(* Logix 5000 project; controller WED2413001_BI600_AB vendor 1 type 14 code 192 rev 35.11; software revision 35.01 *)
// WED2413001_BI600_AB- automatically dispenses film on a roll, cuts, seals and inserts bags into cases, trays and bins

TASK MainTask (continuous, watchdog 500 ms) : BI600_MainProgram

MODULES
   Local : vendor 1 type 14 code 192 (5069 0, rev 35.11)
      VFD1_FILM_UNWIND : PowerFlex 525-EENET (Ethernet 192.168.5.38, rev 7.1, Output RPI 20 ms)   // PowerFlex 525 AC Drive, with Embedded EtherNet/IP and Safety, 200...240V AC, 3 Phase, 5.0 Amps, 1 H
      Cuffer_servo_UpDown : vendor 1 type 37 code 73 (Ethernet 192.168.5.30, rev 13.1, A_MotionDiagnostics RPI 1 ms, B_MotionSync RPI 1 ms)   // ALLEN BRADLEY 2198-C1015-ERS KINETIX 5300 SERVO VARIATEUR, 1.5KW 200V
      Cuffer_servomotor_OpenClose : 2198-C1004-ERS (Ethernet 192.168.5.31, rev 13.1, A_MotionDiagnostics RPI 1 ms, B_MotionSync RPI 1 ms)   // KINETIX 5300 SERVO VARIA TEUR 0.4KW 200V
      SD3_INFEED_CONVEYOR_FRONT : 2198-C1004-ERS (Ethernet 192.168.5.32, rev 13.1, A_MotionDiagnostics RPI 1 ms, B_MotionSync RPI 1 ms)   // KINETIX 5300 SERVO VARIA TEUR 0.4KW 200V
      SD4_INFEED_CONVEYOR_REAR : 2198-C1004-ERS (Ethernet 192.168.5.33, rev 13.1, A_MotionDiagnostics RPI 1 ms, B_MotionSync RPI 1 ms)   // KINETIX 5300 SERVO VARIA TEUR 0.4KW 200V
      SD5_PROCESS_CONVEYOR_FRONT : 2198-C1004-ERS (Ethernet 192.168.5.34, rev 13.1, A_MotionDiagnostics RPI 1 ms, B_MotionSync RPI 1 ms)   // KINETIX 5300 SERVO VARIA TEUR 0.4KW 200V
      SD6_PROCESS_CONVEYOR_REAR : 2198-C1004-ERS (Ethernet 192.168.5.35, rev 13.1, A_MotionDiagnostics RPI 1 ms, B_MotionSync RPI 1 ms)   // KINETIX 5300 SERVO VARIA TEUR 0.4KW 200V
      SD7_SERVO_SEALER_UPDOWN : 2198-C1004-ERS (Ethernet 192.168.5.36, rev 13.1, A_MotionDiagnostics RPI 1 ms, B_MotionSync RPI 1 ms)   // KINETIX 5300 SERVO VARIA TEUR 0.4KW 200V
      SD8_SERVO_FILM_FEED : 2198-C1004-ERS (Ethernet 192.168.5.37, rev 13.1, A_MotionDiagnostics RPI 1 ms, B_MotionSync RPI 1 ms)   // KINETIX 5300 SERVO VARIA TEUR 0.4KW 200V
      EX260SEN2_A : vendor 7 type 27 code 157 (Ethernet 192.168.5.40, rev 1.1, Output RPI 10 ms)   // EX260-SEN2 ETHERNET/IP, NPN (32OUT)
      EX260SEN2_B : vendor 7 type 27 code 157 (Ethernet 192.168.5.41, rev 1.1, Output RPI 10 ms)   // EX260-SEN2 ETHERNET/IP, NPN (32OUT)
      EX260SEN2_C : vendor 7 type 27 code 157 (Ethernet 192.168.5.42, rev 1.1, Output RPI 10 ms)   // EX260-SEN2 ETHERNET/IP, NPN (32OUT)
      EX260SEN2_D : vendor 7 type 27 code 157 (Ethernet 192.168.5.43, rev 1.1, Output RPI 10 ms)   // EX260-SEN2 ETHERNET/IP, NPN (32OUT)
      PLC_INPUTS_2 : 5069-IB16 (5069 2, rev 2.1, StandardDataDriven RPI 5 ms)   // 16 INPUTS
           Local:2:I.Pt00.Data   // RACK 1 SLOT 2 INPUT 0
           Local:2:I.Pt01.Data   // RACK 1 SLOT 2 INPUT 1
           Local:2:I.Pt02.Data   // RACK 1 SLOT 2 INPUT 2
           Local:2:I.Pt03.Data   // RACK 1 SLOT 2 INPUT 3
           Local:2:I.Pt04.Data   // RACK 1 SLOT 2 INPUT 4
           Local:2:I.Pt05.Data   // RACK 1 SLOT 2 INPUT 5
           Local:2:I.Pt06.Data   // RACK 1 SLOT 2 INPUT 6
           Local:2:I.Pt07.Data   // RACK 1 SLOT 2 INPUT 7
           Local:2:I.Pt08.Data   // RACK 1 SLOT 2 INPUT 8
           Local:2:I.Pt09.Data   // RACK 1 SLOT 2 INPUT 9
           Local:2:I.Pt10.Data   // RACK 1 SLOT 2 INPUT 10
           Local:2:I.Pt11.Data   // RACK 1 SLOT 2 INPUT 11
           Local:2:I.Pt12.Data   // RACK 1 SLOT 2 INPUT 12
           Local:2:I.Pt13.Data   // RACK 1 SLOT 2 INPUT 13
           Local:2:I.Pt14.Data   // RACK 1 SLOT 2 INPUT 14
           Local:2:I.Pt15.Data   // RACK 1 SLOT 2 INPUT 15
      PLC_INPUTS_1 : 5069-IB16 (5069 1, rev 2.1, StandardDataDriven RPI 5 ms)   // 16 INPUTS
           Local:1:I.Pt01.Data   // RACK 1 SLOT 1 INPUT 1
           Local:1:I.Pt00.Data   // RACK 1 SLOT 1 INPUT 0
           Local:1:I.Pt02.Data   // RACK 1 SLOT 1 INPUT 2
           Local:1:I.Pt03.Data   // RACK 1 SLOT 1 INPUT 3
           Local:1:I.Pt04.Data   // RACK 1 SLOT 1 INPUT 4
           Local:1:I.Pt05.Data   // RACK 1 SLOT 1 INPUT 5
           Local:1:I.Pt06.Data   // RACK 1 SLOT 1 INPUT 6
           Local:1:I.Pt07.Data   // RACK 1 SLOT 1 INPUT 7
           Local:1:I.Pt08.Data   // RACK 1 SLOT 1 INPUT 8
           Local:1:I.Pt09.Data   // RACK 1 SLOT 1 INPUT 9
           Local:1:I.Pt10.Data   // RACK 1 SLOT 1 INPUT 10
           Local:1:I.Pt11.Data   // RACK 1 SLOT 1 INPUT 11
           Local:1:I.Pt12.Data   // RACK 1 SLOT 1 INPUT 12
           Local:1:I.Pt13.Data   // RACK 1 SLOT 1 INPUT 13
           Local:1:I.Pt14.Data   // RACK 1 SLOT 1 INPUT 14
           Local:1:I.Pt15.Data   // RACK 1 SLOT 1 INPUT 15
      PLC_OUTPUTS_2 : 5069-OB16 (5069 4, rev 3.1, StandardDataDriven RPI 5 ms)   // 16 OUTPUTS
      PLC_OUTPUTS_1 : 5069-OB16 (5069 3, rev 3.1, StandardDataDriven RPI 5 ms)   // 16 OUTPUTS
      PIREG_SEALER : vendor 1547 type 43 code 100 (Ethernet 192.168.5.50, rev 2.1, StandardDataDriven RPI 10 ms)   // These interfaces can be used to control all the controller functions and poll controller information. The ACTUAL temperature of the heat sealing band is supplied to the Analog or EtherNet/IP™ interface as well as to an analog 0 to 10V DC output. The real heat sealing band temperature can thus be displayed on an external temperature meter.
      UNWIND_ENCODER : vendor 1 type 34 code 3 (Ethernet 192.168.5.23, rev 1.1, StandardDataDriven RPI 20 ms)   // UNWIND_ENCODER
END_MODULES

ADD_ON_INSTRUCTION SCP   (* revision 1.2, vendor Rockwell Automation *)
// Scale w/Parameters
// Help:
// Use this instruction to scale data from your analog module and bring it into the limits prescribed by the process variable or another analog module.
// Equations used in calculating a linear relationship:
// Scaled value = (input value - input min.) x rate + scaled minimum
// Rate = (scaled max. - scaled min.) / (input max. - input min.)
VAR_INPUT
   Input : REAL; {required}
   Input_Min : REAL; {required}
   Input_Max : REAL; {required}
   Scaled_Min : REAL; {required}
   Scaled_Max : REAL; {required}
END_VAR
VAR_OUTPUT
   Output : REAL; {access Read Only, required}
END_VAR
VAR
   Rate : REAL;
END_VAR

ROUTINE Logic   (* ladder *)
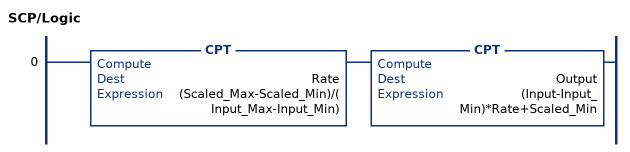
   0: CPT(Rate,(Scaled_Max-Scaled_Min)/(Input_Max-Input_Min))CPT(Output,(Input-Input_Min)*Rate+Scaled_Min);
END_ROUTINE
END_ADD_ON_INSTRUCTION

VAR_GLOBAL   (* controller tags *)
   Action_000 : SFC_ACTION := (Status := 16#0020_0000, PauseTimer := 1);
   Action_001 : SFC_ACTION := (Status := 16#0020_0000, PauseTimer := 1);
   Action_002 : SFC_ACTION := (Status := 16#0020_0000, PauseTimer := 1);
   Action_003 : SFC_ACTION := (Status := 16#0020_0000, PauseTimer := 1);
   Action_004 : SFC_ACTION := (Status := 16#0020_0000, PauseTimer := 1);
   Action_005 : SFC_ACTION := (Status := 16#0020_0000, PauseTimer := 1);
   Action_006 : SFC_ACTION := (Status := 16#0020_0000, PauseTimer := 1);
   Action_007 : SFC_ACTION := (Status := 16#0020_0000, PauseTimer := 1);
   Action_008 : SFC_ACTION := (Status := 16#0020_0000, PauseTimer := 1);
   Action_009 : SFC_ACTION := (Status := 16#0020_0000, PauseTimer := 1);
   Action_010 : SFC_ACTION := (Status := 16#0020_0000, PauseTimer := 1);
   Action_011 : SFC_ACTION := (Status := 16#0020_0000, PauseTimer := 1);
   Action_012 : SFC_ACTION := (Status := 16#0020_0000, PauseTimer := 1);
   Action_013 : SFC_ACTION := (Status := 16#0020_0000, PauseTimer := 1);
   Action_014 : SFC_ACTION := (Status := 16#0020_0000, PauseTimer := 1);
   Action_015 : SFC_ACTION := (Status := 16#0020_0000, PauseTimer := 1);
   Action_016 : SFC_ACTION := (Status := 16#0020_0000, PauseTimer := 1);
   Action_017 : SFC_ACTION := (Status := 16#0020_0000, PauseTimer := 1);
   Action_018 : SFC_ACTION := (Status := 16#0020_0000, PauseTimer := 1);
   Action_019 : SFC_ACTION := (Status := 16#0020_0000, PauseTimer := 1);
   Action_020 : SFC_ACTION := (Status := 16#0020_0000, PauseTimer := 1);
   AIR_PRESSURE_SENSOR : BOOL;
   Always_False : BOOL;
   AXIS_SD1 : AXIS_CIP_DRIVE;
   AXIS_SD2 : AXIS_CIP_DRIVE;
   AXIS_SD3 : AXIS_CIP_DRIVE;
   AXIS_SD4 : AXIS_CIP_DRIVE;
   AXIS_SD5 : AXIS_CIP_DRIVE;
   AXIS_SD6 : AXIS_CIP_DRIVE;
   AXIS_SD7 : AXIS_CIP_DRIVE;
   AXIS_SD8 : AXIS_CIP_DRIVE;
   bBadBagInsert : BOOL;
   C_STOP_BUTTON : BOOL;
   CONTAINER_AT_INFEED : BOOL;
   DANCER_ROLL_DOWN : BOOL;
   DANCER_ROLL_MID : BOOL;
   DANCER_ROLL_OUT_FILM : BOOL;
   DANCER_ROLL_UP : BOOL;
   Delay_ExtendFingers_UP : BOOL;
   Delay_RotateFingers_Up_UP : BOOL;
   DM1_FUNCTION_BUTTON : BOOL;
   DOOR_SS1 : BOOL;
   DOOR_SS2 : BOOL;
   DOOR_SS3 : BOOL;
   DOOR_SS4 : BOOL;
   E_STOP : BOOL;
   E_STOP_PBE1 : BOOL;
   E_STOP_PBE2 : BOOL;
   Enable_Full_FilmFeed : BOOL;
   EXECUTING : BOOL;
   Fast_Init : BOOL;
   First_Scan_Bit : BOOL;
   FixOverShooting : SFC_STEP := (Status := 16#0020_0000, PauseTimer := 1);
   FixOverShooting_Done : SFC_STEP := (Status := 16#0020_0000, PauseTimer := 1);
   Force_Init : BOOL;
   Group_SD : MOTION_GROUP;
   HMI_BoxPassThroughModeEnable : BOOL;
   HMI_Enable_SimMode_Btn : BOOL;
   HOLD_CMD : BOOL;
   InfeedBelt_BoxPassThroug_h_Done : SFC_STEP := (Status := 16#0020_0000, PauseTimer := 1);
   InfeedBelt_BoxPassThroug_h_Running : SFC_STEP := (Status := 16#0020_0000, PauseTimer := 1);
   InfeedBelt_Full : SFC_STEP := (Status := 16#0020_0000, PauseTimer := 1);
   InfeedBelt_Full_Flag : BOOL;
   InfeedBelt_Init : SFC_STEP := (Status := 16#0020_0000, PauseTimer := 1);
   InfeedBelt_PowerON_Status : BOOL;
   InfeedBelt_Run : SFC_STEP := (Status := 16#0020_0000, PauseTimer := 1);
   InfeedBelt_Stop : SFC_STEP := (Status := 16#0020_0000, PauseTimer := 1);
   InfeedBelt_Wait : SFC_STEP := (Status := 16#0020_0000, PauseTimer := 1);
   INFLATOR : BOOL;
   INIT : BOOL;
   Init_Servo_Power_On : BOOL;
   Init_Timer : TIMER;
   INTER_ROLLER : BOOL;
   Machine_State : DINT;
   Master_RESET : BOOL;
   MC_CufferOC_AxisUse_Done : BOOL;
   MC_CufferOC_Pwr_Status : BOOL;
   MC_CufferUD_Axis_to_Unuse_Done : BOOL;
   MC_CufferUD_AxisUse_Done : BOOL;
   MC_CufferUD_Pwr_Status : BOOL;
   MC_FilmFeed_Axis_to_Unuse_Done : BOOL;
   MC_FilmFeed_AxisUse_Done : BOOL;
   MC_FilmFeed_Pwr_Status : BOOL;
   MC_InfeedBelt_Details_Idle : BOOL;
   MC_InfeedBelt_Status_Ready : BOOL;
   MC_MoveABS_CufferOC_Open_Done : BOOL;
   MC_MoveVelocity_InfeedBelt_Busy : BOOL;
   MC_ProcessBelt_ClearConveyr_Done : BOOL;
   MC_SealerUD_Axis_to_Unuse_Done : BOOL;
   MC_SealerUD_AxisUse_Done : BOOL;
   MC_SealerUD_Pwr_Status : BOOL;
   MC_Stop_InfeedBelt_Busy : BOOL;
   MC_Write_CufferOC_Done : BOOL;
   MC_Write_CufferUD_Done : BOOL;
   MC_Write_FilmFeed_Done : BOOL;
   MC_Write_SealerUD_Done : BOOL;
   mInfeedBelt_MC_AxisToUnuse_Done : BOOL;
   mInfeedBelt_MC_AxisToUse_Done : BOOL;
   mInfeedBelt_MC_WritePar_Done : BOOL;
   mMC_CufferUD_ParkPos_Done : BOOL;
   mMC_CufferUD_ParkPos_OverTorqueFix_Done : BOOL;
   mMC_SealerUD_ParkPos_Done : BOOL;
   mProcessBelt_MC_AxisToUnuse_Done : BOOL;
   mProcessBelt_MC_AxisToUse_Done : BOOL;
   mProcessBelt_MC_WritePar_Done : BOOL;
   nfeedBelt_Srv_Geared : BOOL;
   OUTFEED_BACKUP : BOOL;
   Pending_Init : BOOL;
   PHO1 : BOOL;
   Power_ON : BOOL;
   ProcessBelt_Init : SFC_STEP := (Status := 16#0020_0000, PauseTimer := 1);
   ProcessBelt_PowerON_Status : BOOL;
   ProcessBelt_Srv_Geared : BOOL;
   ProcessBelt_Wait : SFC_STEP := (Status := 16#0020_0000, PauseTimer := 1);
   PRODUCTION_CNT : BOOL;
   R00ABORTED : SFC_STEP := (Status := 16#0020_0000, PauseTimer := 1);
   R00ABORTING : SFC_STEP := (Status := 16#0020_0000, PauseTimer := 1);
   R00CLEARING : SFC_STEP := (Status := 16#0020_0000, PauseTimer := 1);
   R00COMPLETE : SFC_STEP := (Status := 16#0020_0000, PauseTimer := 1);
   R00COMPLETING : SFC_STEP := (Status := 16#0020_0000, PauseTimer := 1);
   R00EXECUTE : SFC_STEP := (Status := 16#0020_0000, PauseTimer := 1);
   R00HELD : SFC_STEP := (Status := 16#0020_0000, PauseTimer := 1);
   R00HOLDING : SFC_STEP := (Status := 16#0020_0000, PauseTimer := 1);
   R00IDLE : SFC_STEP := (Status := 16#0020_0000, PauseTimer := 1);
   R00INITIAL : SFC_STEP := (Status := 16#0020_0000, PauseTimer := 1);
   R00RESETING : SFC_STEP := (Status := 16#0020_0000, PauseTimer := 1);
   R00STARTING : SFC_STEP := (Status := 16#0020_0000, PauseTimer := 1);
   R00STOPPED : SFC_STEP := (Status := 16#0020_0000, PauseTimer := 1);
   R00STOPPING : SFC_STEP := (Status := 16#0020_0000, PauseTimer := 1);
   R00SUSPENDED : SFC_STEP := (Status := 16#0020_0000, PauseTimer := 1);
   R00SUSPENDING : SFC_STEP := (Status := 16#0020_0000, PauseTimer := 1);
   R00UNHOLDING : SFC_STEP := (Status := 16#0020_0000, PauseTimer := 1);
   R00UNSUSPENDED : SFC_STEP := (Status := 16#0020_0000, PauseTimer := 1);
   R02_INIT : SFC_STEP := (Status := 16#0020_0000, PauseTimer := 1);
   R02_Init_Clear_Process_Conveyr : SFC_STEP := (Status := 16#0020_0000, PauseTimer := 1);
   R02_Init_CufferUD_To_Park_Pos : SFC_STEP := (Status := 16#0020_0000, PauseTimer := 1);
   R02_Init_Force_ExtendFingers : SFC_STEP := (Status := 16#0020_0000, PauseTimer := 1);
   R02_Init_ForceFingers_UP : SFC_STEP := (Status := 16#0020_0000, PauseTimer := 1);
   R02_Init_GearMotors : SFC_STEP := (Status := 16#0020_0000, PauseTimer := 1);
   R02_Init_MC_Set_Servo_Power : SFC_STEP := (Status := 16#0020_0000, PauseTimer := 1);
   R02_Init_Open_CufferOC : SFC_STEP := (Status := 16#0020_0000, PauseTimer := 1);
   R02_Init_SealerUD_To_Park_Pos : SFC_STEP := (Status := 16#0020_0000, PauseTimer := 1);
   R02_Init_Set_Axis_To_Unused : SFC_STEP := (Status := 16#0020_0000, PauseTimer := 1);
   R02_Init_Set_Axis_To_Used : SFC_STEP := (Status := 16#0020_0000, PauseTimer := 1);
   R02_Init_TOSS : SFC_STEP := (Status := 16#0020_0000, PauseTimer := 1);
   R02_INIT_WAIT : SFC_STEP := (Status := 16#0020_0000, PauseTimer := 1);
   R02_Init_Write_Servo_Params : SFC_STEP := (Status := 16#0020_0000, PauseTimer := 1);
   RESET_CMD : BOOL;
   RESUME_CMD : BOOL;
   SAFETY_CLEAR : BOOL;
   SAFETY_RELAY_SR1 : BOOL;
   SD1_HOME_POSITION : BOOL;
   SH_TEST_DINT : DINT;
   SimulationFlag : BOOL;
   SkipWriteServoPar : BOOL;
   SOLA1_SEALER_JAW : BOOL;
   SOLA2_FILM_NIPROLL_ROLLERS : BOOL;
   SOLA3_KNIFE_SEALING_KNIFE : BOOL;
   SOLB1_FINGERS_DOWN_BACKSIDE : BOOL;
   SOLB2_BACK_PINCH_FINGER_STOPPER : BOOL;
   SOLB3_BACK_FINGERS_OUT : BOOL;
   SOLB4_BACK_RETRACT_SUCTION_CUPS_OUT : BOOL;
   SOLC1_FINGERS_DOWN_FRONTSID : BOOL;
   SOLC2_FRONT_PINCH_FINGER_STOPPER : BOOL;
   SOLC3_FRONT_FINGERS_OUT : BOOL;
   SOLC4_FRONT_RETRACT_SUCTION_CUPS_OUT : BOOL;
   SPARE_SLOT1_INPUT6 : BOOL;
   SPARE_SLOT2_INPUT10 : BOOL;
   SPARE_SLOT2_INPUT11 : BOOL;
   SPARE_SLOT2_INPUT12 : BOOL;
   SPARE_SLOT2_INPUT13 : BOOL;
   SPARE_SLOT2_INPUT14 : BOOL;
   SPARE_SLOT2_INPUT15 : BOOL;
   SPARE_SLOT2_INPUT2 : BOOL;
   SPARE_SLOT2_INPUT4 : BOOL;
   SPARE_SLOT2_INPUT6 : BOOL;
   SPARE_SLOT2_INPUT7 : BOOL;
   SPARE_SLOT2_INPUT8 : BOOL;
   SPARE_SLOT2_INPUT9 : BOOL;
   SPARE_SLOT3_OUTPUT0 : BOOL;
   SPARE_SLOT3_OUTPUT1 : BOOL;
   SPARE_SLOT3_OUTPUT10 : BOOL;
   SPARE_SLOT3_OUTPUT2 : BOOL;
   SPARE_SLOT3_OUTPUT4 : BOOL;
   SPARE_SLOT3_OUTPUT5 : BOOL;
   SPARE_SLOT3_OUTPUT7 : BOOL;
   SPARE_SLOT3_OUTPUT9 : BOOL;
   SPARE_SLOT4_OUTPUT0 : BOOL;
   SPARE_SLOT4_OUTPUT1 : BOOL;
   SPARE_SLOT4_OUTPUT10 : BOOL;
   SPARE_SLOT4_OUTPUT11 : BOOL;
   SPARE_SLOT4_OUTPUT12 : BOOL;
   SPARE_SLOT4_OUTPUT13 : BOOL;
   SPARE_SLOT4_OUTPUT14 : BOOL;
   SPARE_SLOT4_OUTPUT15 : BOOL;
   SPARE_SLOT4_OUTPUT2 : BOOL;
   SPARE_SLOT4_OUTPUT3 : BOOL;
   SPARE_SLOT4_OUTPUT4 : BOOL;
   SPARE_SLOT4_OUTPUT5 : BOOL;
   SPARE_SLOT4_OUTPUT6 : BOOL;
   SPARE_SLOT4_OUTPUT7 : BOOL;
   SPARE_SLOT4_OUTPUT8 : BOOL;
   SPARE_SLOT4_OUTPUT9 : BOOL;
   STACK_LIGHT_BLUE : BOOL;
   STACK_LIGHT_BUZZER : BOOL;
   STACK_LIGHT_GREEN : BOOL;
   STACK_LIGHT_RED : BOOL;
   STACK_LIGHT_WHITE : BOOL;
   START_CMD : BOOL;
   State_Initializing : BOOL;
   State_Running : BOOL;
   State_Stopping : BOOL;
   STOP_CMD : BOOL;
   SUCTION_CUPS_VACUUM : BOOL;
   SUSPEND_CMD : BOOL;
   System_Ready : BOOL;
   TOSS_Connected : BOOL;
   TOSS_Init_Done : BOOL;
   Tran_000 : BOOL;
   Tran_001 : BOOL;
   Tran_002 : BOOL;
   Tran_003 : BOOL;
   Tran_005 : BOOL;
   Tran_006 : BOOL;
   Tran_007 : BOOL;
   Tran_008 : BOOL;
   Tran_009 : BOOL;
   Tran_010 : BOOL;
   Tran_011 : BOOL;
   Tran_012 : BOOL;
   Tran_013 : BOOL;
   Tran_014 : BOOL;
   Tran_015 : BOOL;
   Tran_016 : BOOL;
   Tran_017 : BOOL;
   Tran_018 : BOOL;
   Tran_019 : BOOL;
   Tran_020 : BOOL;
   Tran_021 : BOOL;
   Tran_022 : BOOL;
   Tran_023 : BOOL;
   Tran_024 : BOOL;
   Tran_025 : BOOL;
   Tran_026 : BOOL;
   Tran_027 : BOOL;
   Tran_028 : BOOL;
   Tran_029 : BOOL;
   Tran_030 : BOOL;
   Tran_031 : BOOL;
   Tran_032 : BOOL;
   Tran_033 : BOOL;
   Tran_034 : BOOL;
   Tran_035 : BOOL;
   Tran_036 : BOOL;
   Tran_037 : BOOL;
   Tran_038 : BOOL;
   Tran_039 : BOOL;
   Tran_040 : BOOL;
   Tran_041 : BOOL;
   Tran_042 : BOOL;
   Tran_043 : BOOL;
   Tran_044 : BOOL;
   Tran_045 : BOOL;
   Tran_046 : BOOL;
   UNWIND_DOOR_SS : BOOL;
   Vacuum_ON : BOOL;
   VACUUM_SWITCH : BOOL;
END_VAR

PROGRAM BI600_MainProgram   (* main routine R00_Main *)

ROUTINE R001_Inputs   (* ladder *)
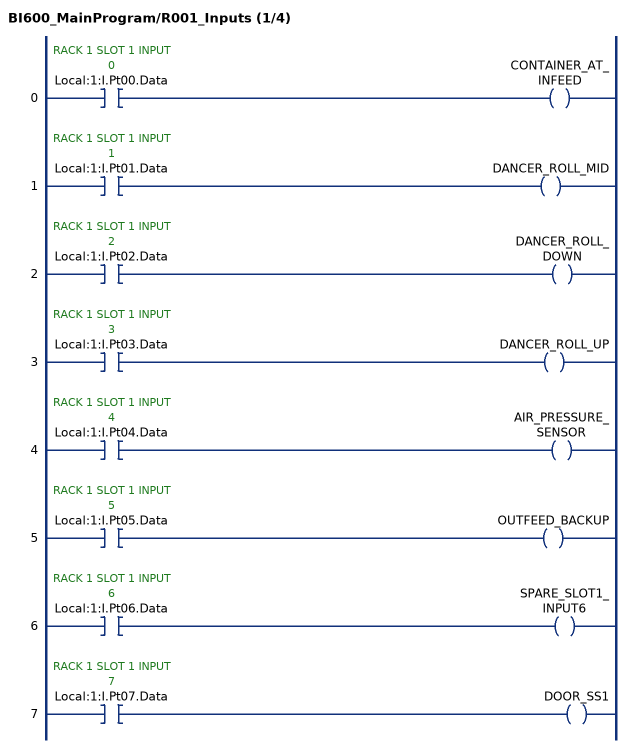
   0: XIC(Local:1:I.Pt00.Data)OTE(CONTAINER_AT_INFEED);
   1: XIC(Local:1:I.Pt01.Data)OTE(DANCER_ROLL_MID);
   2: XIC(Local:1:I.Pt02.Data)OTE(DANCER_ROLL_DOWN);
   3: XIC(Local:1:I.Pt03.Data)OTE(DANCER_ROLL_UP);
   4: XIC(Local:1:I.Pt04.Data)OTE(AIR_PRESSURE_SENSOR);
   5: XIC(Local:1:I.Pt05.Data)OTE(OUTFEED_BACKUP);
   6: XIC(Local:1:I.Pt06.Data)OTE(SPARE_SLOT1_INPUT6);
   7: XIC(Local:1:I.Pt07.Data)OTE(DOOR_SS1);
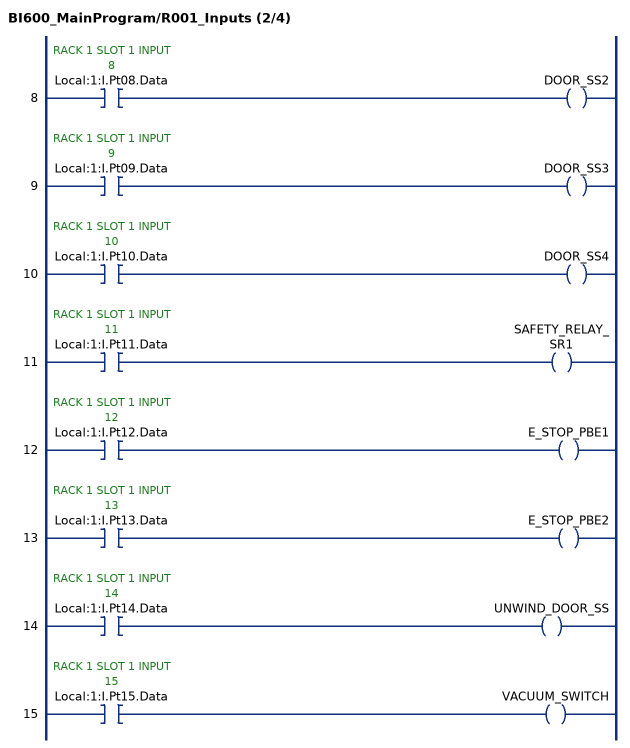
   8: XIC(Local:1:I.Pt08.Data)OTE(DOOR_SS2);
   9: XIC(Local:1:I.Pt09.Data)OTE(DOOR_SS3);
   10: XIC(Local:1:I.Pt10.Data)OTE(DOOR_SS4);
   11: XIC(Local:1:I.Pt11.Data)OTE(SAFETY_RELAY_SR1);
   12: XIC(Local:1:I.Pt12.Data)OTE(E_STOP_PBE1);
   13: XIC(Local:1:I.Pt13.Data)OTE(E_STOP_PBE2);
   14: XIC(Local:1:I.Pt14.Data)OTE(UNWIND_DOOR_SS);
   15: XIC(Local:1:I.Pt15.Data)OTE(VACUUM_SWITCH);
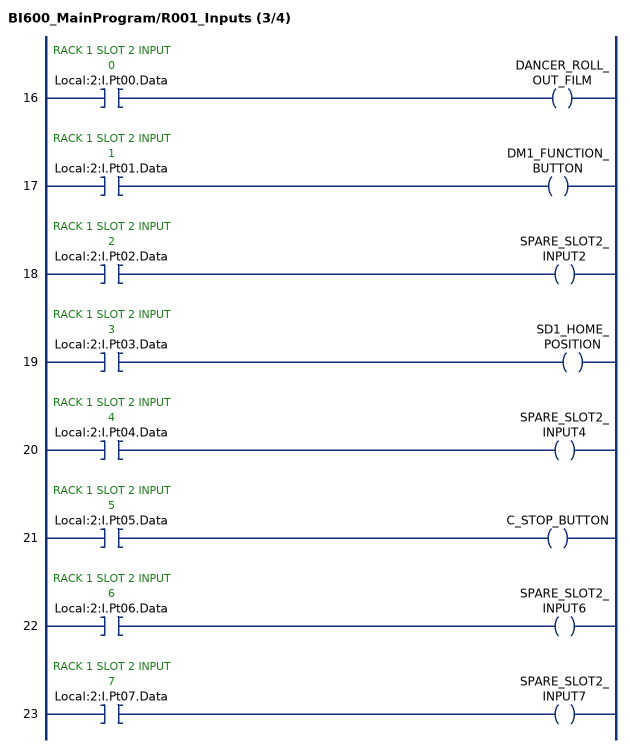
   16: XIC(Local:2:I.Pt00.Data)OTE(DANCER_ROLL_OUT_FILM);
   17: XIC(Local:2:I.Pt01.Data)OTE(DM1_FUNCTION_BUTTON);
   18: XIC(Local:2:I.Pt02.Data)OTE(SPARE_SLOT2_INPUT2);
   19: XIC(Local:2:I.Pt03.Data)OTE(SD1_HOME_POSITION);
   20: XIC(Local:2:I.Pt04.Data)OTE(SPARE_SLOT2_INPUT4);
   21: XIC(Local:2:I.Pt05.Data)OTE(C_STOP_BUTTON);
   22: XIC(Local:2:I.Pt06.Data)OTE(SPARE_SLOT2_INPUT6);
   23: XIC(Local:2:I.Pt07.Data)OTE(SPARE_SLOT2_INPUT7);
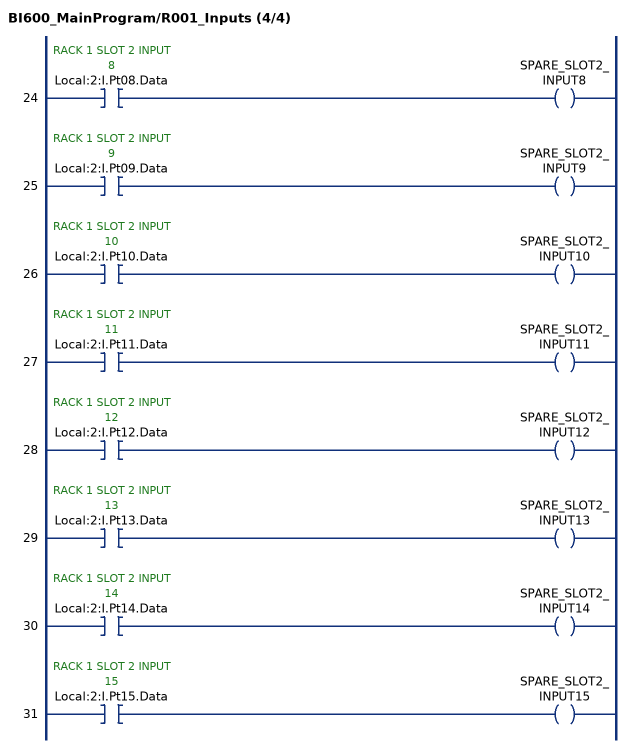
   24: XIC(Local:2:I.Pt08.Data)OTE(SPARE_SLOT2_INPUT8);
   25: XIC(Local:2:I.Pt09.Data)OTE(SPARE_SLOT2_INPUT9);
   26: XIC(Local:2:I.Pt10.Data)OTE(SPARE_SLOT2_INPUT10);
   27: XIC(Local:2:I.Pt11.Data)OTE(SPARE_SLOT2_INPUT11);
   28: XIC(Local:2:I.Pt12.Data)OTE(SPARE_SLOT2_INPUT12);
   29: XIC(Local:2:I.Pt13.Data)OTE(SPARE_SLOT2_INPUT13);
   30: XIC(Local:2:I.Pt14.Data)OTE(SPARE_SLOT2_INPUT14);
   31: XIC(Local:2:I.Pt15.Data)OTE(SPARE_SLOT2_INPUT15);
END_ROUTINE

ROUTINE R00_Machine_Mode_State   (* ladder *)
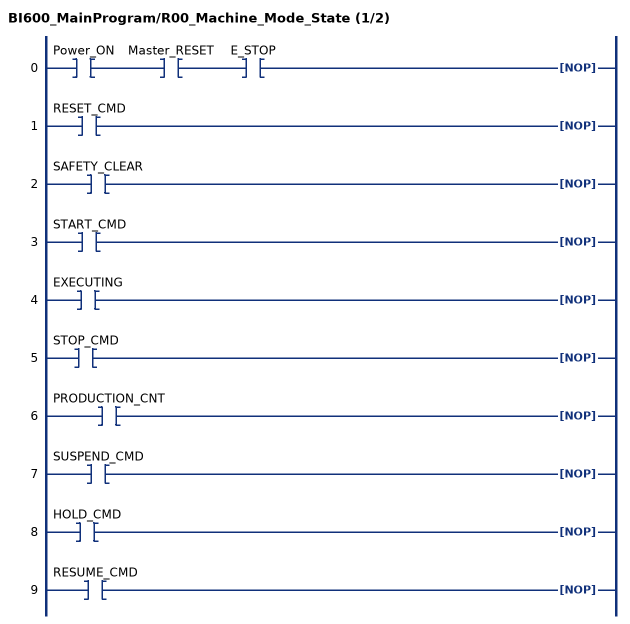
   0: XIC(Power_ON)XIC(Master_RESET)XIC(E_STOP)NOP();
   1: XIC(RESET_CMD)NOP();
   2: XIC(SAFETY_CLEAR)NOP();
   3: XIC(START_CMD)NOP();
   4: XIC(EXECUTING)NOP();
   5: XIC(STOP_CMD)NOP();
   6: XIC(PRODUCTION_CNT)NOP();
   7: XIC(SUSPEND_CMD)NOP();
   8: XIC(HOLD_CMD)NOP();
   9: XIC(RESUME_CMD)NOP();
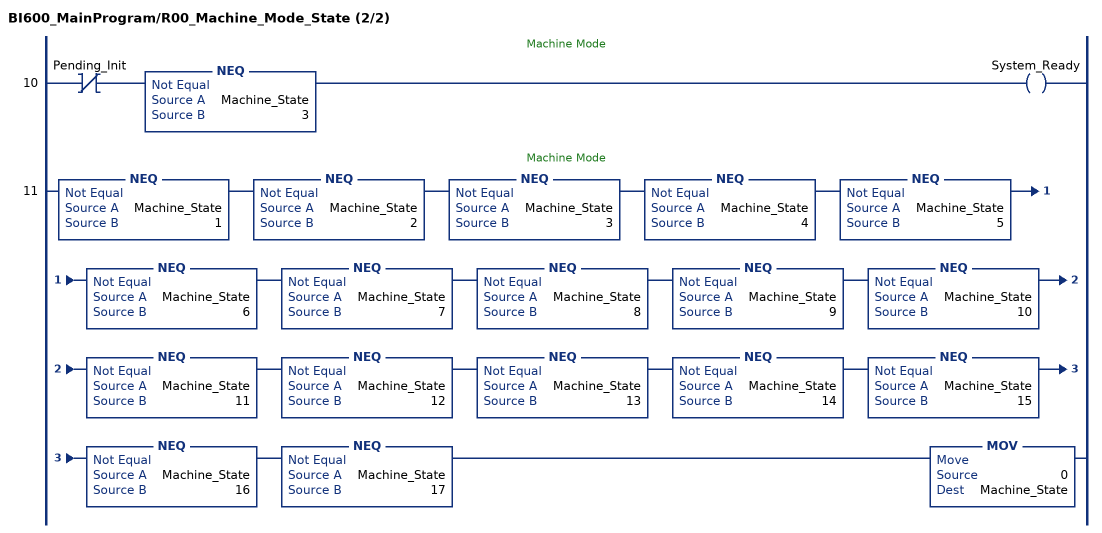
   // Machine Mode
   10: XIO(Pending_Init)NEQ(Machine_State,3)OTE(System_Ready);
   // Machine Mode
   11: NEQ(Machine_State,1)NEQ(Machine_State,2)NEQ(Machine_State,3)NEQ(Machine_State,4)NEQ(Machine_State,5)NEQ(Machine_State,6)NEQ(Machine_State,7)NEQ(Machine_State,8)NEQ(Machine_State,9)NEQ(Machine_State,10)NEQ(Machine_State,11)NEQ(Machine_State,12)NEQ(Machine_State,13)NEQ(Machine_State,14)NEQ(Machine_State,15)NEQ(Machine_State,16)NEQ(Machine_State,17)MOV(0,Machine_State);
END_ROUTINE

ROUTINE R00_Machine_Mode_StateSFC   (* sequential function chart *)